
PopupScreen "Tank 1S Status" 480x272
   TextField "Text field_4" at 9,135 size 86x22; Text 'Pressure:'
   IOField "I/O field_1" at 139,130 size 90x25; FormatPattern s999.9; Unit  mBar
      ProcessValue <- "20_TANKS_IP_DATA_RIO_01_THIRD_TANK_TANKS_PRESS"
   TextField "Text field_5" at 9,169 size 113x22; Text 'Water Level:'
   IOField "I/O field_2" at 138,164 size 90x25; FormatPattern 999.9; Unit  %
      ProcessValue <- "20_TANKS_IP_DATA_RIO_01_THIRD_TANK_BWT_LEVEL"
   TextField "Text field_6" at 9,203 size 137x22; Text 'MBG Flow Rate:'
   IOField "I/O field_3" at 139,198 size 90x25; FormatPattern 999.9; Unit  m³/hr
      ProcessValue <- "20_TANKS_IP_DATA_RIO_01_THIRD_TANK_MBG_FLOW"
   TextField "Text field_7" at 9,237 size 135x22; Text 'USD Flow Rate:'
   IOField "I/O field_4" at 139,232 size 90x25; FormatPattern 999.9; Unit  m³/hr
      ProcessValue <- "20_TANKS_IP_DATA_RIO_01_THIRD_TANK_USD_FLOW"
   Button "Button_1" at 50,5 size 191x35; TextOff 'Starboard Tank 1 (1S)'
      on Release: function_efd93a16("Tank 1S Status", 0, 0, -1, 0, 1)
   TextField "Text field_1" at 4,90 size 109x25; Text 'TIME LEFT:'
   GraphicView "Graphic view_1" at 9,46 size 228x32; Picture "Tank Manually Disabled"
   GraphicIOField "Graphic I/O field_1" at 9,46 size 228x32; PictureList "Tank Process Stage_II"
      ProcessValue <- "2100_BTCS_CNTRL_DB_BTCS_STATE"
      Visibility <- "504_Tank Grouping_DB2020_GROUP of TANK 3"
   Button "Button_2" at 4,5 size 45x35; TextOff 'Text'; PictureOff "Graphic_286"
      on Click: function_efd93a16("Tank 1S Status", 0, 0, -1, -1, 1)
   IOField "I/O field_29" at 190,90 size 47x25; FormatPattern 99; Unit m
      ProcessValue <- "504_Tank Grouping_DB2020_Time Left Tank_Time Left m Tank 3"
   IOField "I/O field_8" at 147,90 size 42x25; FormatPattern 99; Unit h
      ProcessValue <- "504_Tank Grouping_DB2020_Time Left Tank_Time Left h Tank 3"
   IOField "I/O field_9" at 104,90 size 42x25; FormatPattern 99; Unit d
      ProcessValue <- "504_Tank Grouping_DB2020_Time Left Tank_Time Left d Tank 3"
   TextField "Text field_8" at 241,134 size 140x22; Text 'Water pH Level:'
   IOField "I/O field_5" at 383,129 size 90x25; FormatPattern 99.9
      ProcessValue <- "20_TANKS_IP_DATA_RIO_01_THIRD_TANK_BWT_PH"
   TextField "Text field_9" at 242,168 size 143x22; Text 'Water DO Level:'
   IOField "I/O field_6" at 383,163 size 90x25; FormatPattern 99.99; Unit  mg/l
      ProcessValue <- "20_TANKS_IP_DATA_RIO_01_THIRD_TANK_BWT_DO"
   TextField "Text field_10" at 241,202 size 174x22; Text 'Water Temperature:'
   IOField "I/O field_7" at 398,197 size 75x25; FormatPattern 999.9; Unit  °C
      ProcessValue <- "20_TANKS_IP_DATA_RIO_01_THIRD_TANK_BWT_TEMP"
   Button "Button_5" at 249,229 size 223x40; TextOff 'Tank Shutdown Alarm'
      Visibility <- "2062_Warning_Data_Alarm Tank S1"
   Button "Button_6" at 248,229 size 224x40; TextOff 'No/Low Water Level'; Authorization "Operate"
      Visibility <- "LT421 1S  TANK LEVEL ALARM_ALARM L"

PopupScreen "Tank 2S Status" 480x272
   TextField "Text field_4" at 4,134 size 86x22; Text 'Pressure:'
   IOField "I/O field_1" at 147,129 size 90x25; FormatPattern s999.9; Unit  mBar
      ProcessValue <- "20_TANKS_IP_DATA_RIO_02_SECOND_TANK_TANKS_PRESS"
   TextField "Text field_5" at 4,168 size 113x22; Text 'Water Level:'
   IOField "I/O field_2" at 147,163 size 90x25; FormatPattern 999.9; Unit  %
      ProcessValue <- "20_TANKS_IP_DATA_RIO_02_SECOND_TANK_BWT_LEVEL"
   TextField "Text field_6" at 4,202 size 137x22; Text 'MBG Flow Rate:'
   IOField "I/O field_3" at 147,197 size 90x25; FormatPattern 999.9; Unit  m³/hr
      ProcessValue <- "20_TANKS_IP_DATA_RIO_02_SECOND_TANK_MBG_FLOW"
   TextField "Text field_7" at 4,236 size 135x22; Text 'USD Flow Rate:'
   IOField "I/O field_4" at 147,231 size 90x25; FormatPattern 999.9; Unit  m³/hr
      ProcessValue <- "20_TANKS_IP_DATA_RIO_02_SECOND_TANK_USD_FLOW"
   Button "Button_1" at 50,5 size 191x35; TextOff 'Starboard Tank 2 (2S)'
      on Release: function_efd93a16("Tank 2S Status", 0, 0, -1, 0, 1)
   TextField "Text field_1" at 5,90 size 109x25; Text 'TIME LEFT:'
   GraphicView "Graphic view_1" at 9,46 size 225x32; Picture "Tank Manually Disabled"
   GraphicIOField "Graphic I/O field_1" at 9,46 size 227x32; PictureList "Tank Process Stage_II"
      ProcessValue <- "2100_BTCS_CNTRL_DB_BTCS_STATE"
      Visibility <- "504_Tank Grouping_DB2020_GROUP of TANK 5"
   Button "Button_2" at 4,5 size 45x35; TextOff 'Text'; PictureOff "Graphic_286"
      on Click: function_efd93a16("Tank 2S Status", 0, 0, -1, -1, 1)
   IOField "I/O field_29" at 189,89 size 47x25; FormatPattern 99; Unit m
      ProcessValue <- "504_Tank Grouping_DB2020_Time Left Tank_Time Left m Tank 5"
   IOField "I/O field_8" at 146,90 size 42x25; FormatPattern 99; Unit h
      ProcessValue <- "504_Tank Grouping_DB2020_Time Left Tank_Time Left h Tank 5"
   IOField "I/O field_9" at 103,90 size 42x25; FormatPattern 99; Unit d
      ProcessValue <- "504_Tank Grouping_DB2020_Time Left Tank_Time Left d Tank 5"
   TextField "Text field_8" at 243,133 size 140x22; Text 'Water pH Level:'
   IOField "I/O field_5" at 382,128 size 90x25; FormatPattern 99.9
      ProcessValue <- "20_TANKS_IP_DATA_RIO_02_SECOND_TANK_BWT_PH"
   TextField "Text field_9" at 243,167 size 143x22; Text 'Water DO Level:'
   IOField "I/O field_6" at 382,162 size 90x25; FormatPattern 99.99; Unit  mg/l
      ProcessValue <- "20_TANKS_IP_DATA_RIO_02_SECOND_TANK_BWT_DO"
   TextField "Text field_10" at 243,201 size 174x22; Text 'Water Temperature:'
   IOField "I/O field_7" at 397,196 size 75x25; FormatPattern 999.9; Unit  °C
      ProcessValue <- "20_TANKS_IP_DATA_RIO_02_SECOND_TANK_BWT_TEMP"
   Group "Group" at 245,228 size 227x40
   Button "Button_5" at 245,228 size 227x40; TextOff 'Tank Shutdown Alarm'
      Visibility <- "2062_Warning_Data_Alarm Tank S2"
   Button "Button_6" at 245,228 size 227x40; TextOff 'No/Low Water Level'; Authorization "Operate"
      Visibility <- "LT421 2S  TANK LEVEL ALARM_ALARM L"

PopupScreen "Tank 2P Status" 480x272
   TextField "Text field_4" at 8,135 size 86x22; Text 'Pressure:'
   IOField "I/O field_1" at 139,130 size 90x25; FormatPattern s999.9; Unit  mBar
      ProcessValue <- "20_TANKS_IP_DATA_RIO_02_FIRST_TANK_TANKS_PRESS"
   TextField "Text field_5" at 8,169 size 113x22; Text 'Water Level:'
   IOField "I/O field_2" at 139,164 size 90x25; FormatPattern 999.9; Unit  %
      ProcessValue <- "20_TANKS_IP_DATA_RIO_02_FIRST_TANK_BWT_LEVEL"
   TextField "Text field_6" at 8,203 size 137x22; Text 'MBG Flow Rate:'
   IOField "I/O field_3" at 139,198 size 90x25; FormatPattern 999.9; Unit  m³/hr
      ProcessValue <- "20_TANKS_IP_DATA_RIO_02_FIRST_TANK_MBG_FLOW"
   TextField "Text field_7" at 8,237 size 135x22; Text 'USD Flow Rate:'
   IOField "I/O field_4" at 139,232 size 90x25; FormatPattern 999.9; Unit  m³/hr
      ProcessValue <- "20_TANKS_IP_DATA_RIO_02_FIRST_TANK_USD_FLOW"
   Button "Button_1" at 51,5 size 188x35; TextOff 'Port Tank 2 (2P)'
      on Release: function_efd93a16("Tank 2P Status", 0, 0, -1, 0, 1)
   TextField "Text field_1" at 4,90 size 109x25; Text 'TIME LEFT:'
   GraphicView "Graphic view_1" at 9,46 size 225x32; Picture "Tank Manually Disabled"
   GraphicIOField "Graphic I/O field_1" at 9,46 size 225x32; PictureList "Tank Process Stage_II"
      ProcessValue <- "2100_BTCS_CNTRL_DB_BTCS_STATE"
      Visibility <- "504_Tank Grouping_DB2020_GROUP of TANK 4"
   Button "Button_2" at 4,5 size 45x35; TextOff 'Text'; PictureOff "Graphic_286"
      on Click: function_efd93a16("Tank 2P Status", 0, 0, -1, -1, 1)
   IOField "I/O field_29" at 187,90 size 47x25; FormatPattern 99; Unit m
      ProcessValue <- "504_Tank Grouping_DB2020_Time Left Tank_Time Left m Tank 4"
   IOField "I/O field_8" at 144,90 size 42x25; FormatPattern 99; Unit h
      ProcessValue <- "504_Tank Grouping_DB2020_Time Left Tank_Time Left h Tank 4"
   IOField "I/O field_9" at 101,90 size 42x25; FormatPattern 99; Unit d
      ProcessValue <- "504_Tank Grouping_DB2020_Time Left Tank_Time Left d Tank 4"
   TextField "Text field_8" at 245,135 size 140x22; Text 'Water pH Level:'
   IOField "I/O field_5" at 385,130 size 90x25; FormatPattern 99.9
      ProcessValue <- "20_TANKS_IP_DATA_RIO_02_FIRST_TANK_BWT_PH"
   TextField "Text field_9" at 245,169 size 143x22; Text 'Water DO Level:'
   IOField "I/O field_6" at 385,164 size 90x25; FormatPattern 99.99; Unit  mg/l
      ProcessValue <- "20_TANKS_IP_DATA_RIO_02_FIRST_TANK_BWT_DO"
   TextField "Text field_10" at 245,203 size 174x22; Text 'Water Temperature:'
   IOField "I/O field_7" at 400,198 size 75x25; FormatPattern 999.9; Unit  °C
      ProcessValue <- "20_TANKS_IP_DATA_RIO_02_FIRST_TANK_BWT_TEMP"
   Group "Group" at 244,226 size 230x40
   Button "Button_5" at 244,226 size 230x40; TextOff 'Tank Shutdown Alarm'
      Visibility <- "2062_Warning_Data_Alarm Tank P2"
   Button "Button_6" at 244,226 size 230x40; TextOff 'No/Low Water Level'; Authorization "Operate"
      Visibility <- "FIT418_2P_ALM_ANALOG_DB_ALARM L"

PopupScreen "Tank 3S Status" 480x272
   TextField "Text field_4" at 9,135 size 86x22; Text 'Pressure:'
   IOField "I/O field_1" at 146,130 size 90x25; FormatPattern s999.9; Unit  mBar
      ProcessValue <- "20_TANKS_IP_DATA_RIO_03_SECOND_TANK_TANKS_PRESS"
   TextField "Text field_5" at 9,169 size 113x22; Text 'Water Level:'
   IOField "I/O field_2" at 146,164 size 90x25; FormatPattern 999.9; Unit  %
      ProcessValue <- "20_TANKS_IP_DATA_RIO_03_SECOND_TANK_BWT_LEVEL"
   TextField "Text field_6" at 9,203 size 137x22; Text 'MBG Flow Rate:'
   IOField "I/O field_3" at 146,198 size 90x25; FormatPattern 999.9; Unit  m³/hr
      ProcessValue <- "20_TANKS_IP_DATA_RIO_03_SECOND_TANK_MBG_FLOW"
   TextField "Text field_7" at 9,237 size 135x22; Text 'USD Flow Rate:'
   IOField "I/O field_4" at 146,232 size 90x25; FormatPattern 999.9; Unit  m³/hr
      ProcessValue <- "20_TANKS_IP_DATA_RIO_03_SECOND_TANK_USD_FLOW"
   Button "Button_1" at 51,5 size 189x35; TextOff 'Starboard Tank 3 (3S)'
      on Release: function_efd93a16("Tank 3S Status", 0, 0, -1, 0, 1)
   TextField "Text field_1" at 5,90 size 109x25; Text 'TIME LEFT:'
   GraphicView "Graphic view_1" at 9,46 size 226x32; Picture "Tank Manually Disabled"
   GraphicIOField "Graphic I/O field_1" at 9,46 size 226x32; PictureList "Tank Process Stage_II"
      ProcessValue <- "2100_BTCS_CNTRL_DB_BTCS_STATE"
      Visibility <- "504_Tank Grouping_DB2020_GROUP of TANK 7"
   Button "Button_2" at 4,5 size 45x35; TextOff 'Text'; PictureOff "Graphic_286"
      on Click: function_efd93a16("Tank 3S Status", 0, 0, -1, -1, 1)
   IOField "I/O field_29" at 189,90 size 47x25; FormatPattern 99; Unit m
      ProcessValue <- "504_Tank Grouping_DB2020_Time Left Tank_Time Left m Tank 7"
   IOField "I/O field_8" at 146,90 size 42x25; FormatPattern 99; Unit h
      ProcessValue <- "504_Tank Grouping_DB2020_Time Left Tank_Time Left h Tank 7"
   IOField "I/O field_9" at 103,90 size 42x25; FormatPattern 99; Unit d
      ProcessValue <- "504_Tank Grouping_DB2020_Time Left Tank_Time Left d Tank 7"
   TextField "Text field_8" at 243,135 size 140x22; Text 'Water pH Level:'
   IOField "I/O field_5" at 383,130 size 90x25; FormatPattern 99.9
      ProcessValue <- "20_TANKS_IP_DATA_RIO_03_SECOND_TANK_BWT_PH"
   TextField "Text field_9" at 243,169 size 143x22; Text 'Water DO Level:'
   IOField "I/O field_6" at 383,164 size 90x25; FormatPattern 99.99; Unit  mg/l
      ProcessValue <- "20_TANKS_IP_DATA_RIO_03_SECOND_TANK_BWT_DO"
   TextField "Text field_10" at 243,203 size 174x22; Text 'Water Temperature:'
   IOField "I/O field_7" at 398,198 size 75x25; FormatPattern 999.9; Unit  °C
      ProcessValue <- "20_TANKS_IP_DATA_RIO_03_SECOND_TANK_BWT_TEMP"
   Group "Group" at 243,228 size 230x40
   Button "Button_5" at 243,228 size 230x40; TextOff 'Tank Shutdown Alarm'
      Visibility <- "2062_Warning_Data_Alarm Tank S3"
   Button "Button_6" at 243,228 size 230x40; TextOff 'No/Low Water Level'; Authorization "Operate"
      Visibility <- "LT421 3S  TANK LEVEL ALARM_ALARM L"

PopupScreen "Tank 3P Status" 480x272
   TextField "Text field_4" at 10,135 size 86x22; Text 'Pressure:'
   IOField "I/O field_1" at 148,130 size 90x25; FormatPattern s999.9; Unit  mBar
      ProcessValue <- "20_TANKS_IP_DATA_RIO_03_FIRST_TANK_TANKS_PRESS"
   TextField "Text field_5" at 10,169 size 113x22; Text 'Water Level:'
   IOField "I/O field_2" at 148,164 size 90x25; FormatPattern 999.9; Unit  %
      ProcessValue <- "20_TANKS_IP_DATA_RIO_03_FIRST_TANK_BWT_LEVEL"
   TextField "Text field_6" at 10,203 size 137x22; Text 'MBG Flow Rate:'
   IOField "I/O field_3" at 148,198 size 90x25; FormatPattern 999.9; Unit  m³/hr
      ProcessValue <- "20_TANKS_IP_DATA_RIO_03_FIRST_TANK_MBG_FLOW"
   TextField "Text field_7" at 10,237 size 135x22; Text 'USD Flow Rate:'
   IOField "I/O field_4" at 148,232 size 90x25; FormatPattern 999.9; Unit  m³/hr
      ProcessValue <- "20_TANKS_IP_DATA_RIO_03_FIRST_TANK_USD_FLOW"
   Button "Button_1" at 51,5 size 191x35; TextOff 'Port Tank 3 (3P)'
      on Release: function_efd93a16("Tank 3P Status", 0, 0, -1, 0, 1)
   TextField "Text field_1" at 6,90 size 109x25; Text 'TIME LEFT:'
   GraphicView "Graphic view_1" at 9,46 size 228x32; Picture "Tank Manually Disabled"
   GraphicIOField "Graphic I/O field_1" at 9,46 size 228x32; PictureList "Tank Process Stage_II"
      ProcessValue <- "2100_BTCS_CNTRL_DB_BTCS_STATE"
      Visibility <- "504_Tank Grouping_DB2020_GROUP of TANK 6"
   Button "Button_2" at 4,5 size 45x35; TextOff 'Text'; PictureOff "Graphic_286"
      on Click: function_efd93a16("Tank 3P Status", 0, 0, -1, -1, 1)
   IOField "I/O field_29" at 190,90 size 47x25; FormatPattern 99; Unit m
      ProcessValue <- "504_Tank Grouping_DB2020_Time Left Tank_Time Left m Tank 6"
   IOField "I/O field_8" at 147,90 size 42x25; FormatPattern 99; Unit h
      ProcessValue <- "504_Tank Grouping_DB2020_Time Left Tank_Time Left h Tank 6"
   IOField "I/O field_9" at 104,90 size 42x25; FormatPattern 99; Unit d
      ProcessValue <- "504_Tank Grouping_DB2020_Time Left Tank_Time Left d Tank 6"
   TextField "Text field_8" at 244,135 size 140x22; Text 'Water pH Level:'
   IOField "I/O field_5" at 383,130 size 90x25; FormatPattern 99.9
      ProcessValue <- "20_TANKS_IP_DATA_RIO_03_FIRST_TANK_BWT_PH"
   TextField "Text field_9" at 244,169 size 143x22; Text 'Water DO Level:'
   IOField "I/O field_6" at 383,164 size 90x25; FormatPattern 99.99; Unit  mg/l
      ProcessValue <- "20_TANKS_IP_DATA_RIO_03_FIRST_TANK_BWT_DO"
   TextField "Text field_10" at 244,203 size 174x22; Text 'Water Temperature:'
   IOField "I/O field_7" at 398,198 size 75x25; FormatPattern 999.9; Unit  °C
      ProcessValue <- "20_TANKS_IP_DATA_RIO_03_FIRST_TANK_BWT_TEMP"
   Group "Group" at 247,227 size 226x40
   Button "Button_5" at 247,227 size 226x40; TextOff 'Tank Shutdown Alarm'
      Visibility <- "2062_Warning_Data_Alarm Tank P3"
   Button "Button_6" at 247,227 size 226x40; TextOff 'No/Low Water Level'; Authorization "Operate"
      Visibility <- "LT422 3P  TANK LEVEL ALARM_ALARM L"

PopupScreen "Tank 4S Status" 480x272
   TextField "Text field_4" at 9,135 size 86x22; Text 'Pressure:'
   IOField "I/O field_1" at 147,130 size 90x25; FormatPattern s999.9; Unit  mBar
      ProcessValue <- "20_TANKS_IP_DATA_RIO_04_SECOND_TANK_TANKS_PRESS"
   TextField "Text field_5" at 9,169 size 113x22; Text 'Water Level:'
   IOField "I/O field_2" at 147,164 size 90x25; FormatPattern 999.9; Unit  %
      ProcessValue <- "20_TANKS_IP_DATA_RIO_04_SECOND_TANK_BWT_LEVEL"
   TextField "Text field_6" at 9,203 size 137x22; Text 'MBG Flow Rate:'
   IOField "I/O field_3" at 147,198 size 90x25; FormatPattern 999.9; Unit  m³/hr
      ProcessValue <- "20_TANKS_IP_DATA_RIO_04_SECOND_TANK_MBG_FLOW"
   TextField "Text field_7" at 9,237 size 135x22; Text 'USD Flow Rate:'
   IOField "I/O field_4" at 147,232 size 90x25; FormatPattern 999.9; Unit  m³/hr
      ProcessValue <- "20_TANKS_IP_DATA_RIO_04_SECOND_TANK_USD_FLOW"
   Button "Button_1" at 50,5 size 191x35; TextOff 'Starboard Tank 4 (4S)'
      on Release: function_efd93a16("Tank 4S Status", 0, 0, -1, 2, 1)
   TextField "Text field_1" at 5,90 size 109x25; Text 'TIME LEFT:'
   GraphicView "Graphic view_1" at 9,46 size 227x32; Picture "Tank Manually Disabled"
   GraphicIOField "Graphic I/O field_1" at 9,46 size 227x32; PictureList "Tank Process Stage_II"
      ProcessValue <- "2100_BTCS_CNTRL_DB_BTCS_STATE"
      Visibility <- "504_Tank Grouping_DB2020_GROUP of TANK 9"
   Button "Button_2" at 4,5 size 45x35; TextOff 'Text'; PictureOff "Graphic_286"
      on Click: function_efd93a16("Tank 4S Status", 0, 0, -1, -1, 1)
   IOField "I/O field_29" at 189,90 size 47x25; FormatPattern 99; Unit m
      ProcessValue <- "504_Tank Grouping_DB2020_Time Left Tank_Time Left m Tank 9"
   IOField "I/O field_8" at 146,90 size 42x25; FormatPattern 99; Unit h
      ProcessValue <- "504_Tank Grouping_DB2020_Time Left Tank_Time Left h Tank 9"
   IOField "I/O field_9" at 103,90 size 42x25; FormatPattern 99; Unit d
      ProcessValue <- "504_Tank Grouping_DB2020_Time Left Tank_Time Left d Tank 9"
   TextField "Text field_8" at 243,135 size 140x22; Text 'Water pH Level:'
   IOField "I/O field_5" at 383,130 size 90x25; FormatPattern 99.9
      ProcessValue <- "20_TANKS_IP_DATA_RIO_04_SECOND_TANK_BWT_PH"
   TextField "Text field_9" at 243,169 size 143x22; Text 'Water DO Level:'
   IOField "I/O field_6" at 383,164 size 90x25; FormatPattern 99.99; Unit  mg/l
      ProcessValue <- "20_TANKS_IP_DATA_RIO_04_SECOND_TANK_BWT_DO"
   TextField "Text field_10" at 243,203 size 174x22; Text 'Water Temperature:'
   IOField "I/O field_7" at 398,198 size 75x25; FormatPattern 999.9; Unit  °C
      ProcessValue <- "20_TANKS_IP_DATA_RIO_04_SECOND_TANK_BWT_TEMP"
   Group "Group" at 243,227 size 230x40
   Button "Button_5" at 243,227 size 230x40; TextOff 'Tank Shutdown Alarm'
      Visibility <- "2062_Warning_Data_Alarm Tank S4"
   Button "Button_6" at 243,227 size 230x40; TextOff 'No/Low Water Level'; Authorization "Operate"
      Visibility <- "LT421 4S  TANK LEVEL ALARM_ALARM L"

PopupScreen "Tank 4P Status" 480x272
   TextField "Text field_4" at 9,135 size 86x22; Text 'Pressure:'
   IOField "I/O field_1" at 148,130 size 90x25; FormatPattern s999.9; Unit  mBar
      ProcessValue <- "20_TANKS_IP_DATA_RIO_04_FIRST_TANK_TANKS_PRESS"
   TextField "Text field_5" at 9,169 size 113x22; Text 'Water Level:'
   IOField "I/O field_2" at 148,164 size 90x25; FormatPattern 999.9; Unit  %
      ProcessValue <- "20_TANKS_IP_DATA_RIO_04_FIRST_TANK_BWT_LEVEL"
   TextField "Text field_6" at 9,203 size 137x22; Text 'MBG Flow Rate:'
   IOField "I/O field_3" at 148,198 size 90x25; FormatPattern 999.9; Unit  m³/hr
      ProcessValue <- "20_TANKS_IP_DATA_RIO_04_FIRST_TANK_MBG_FLOW"
   TextField "Text field_7" at 9,237 size 135x22; Text 'USD Flow Rate:'
   IOField "I/O field_4" at 148,232 size 90x25; FormatPattern 999.9; Unit  m³/hr
      ProcessValue <- "20_TANKS_IP_DATA_RIO_04_FIRST_TANK_USD_FLOW"
   Button "Button_1" at 51,5 size 191x35; TextOff 'Port Tank 4 (4P)'
      on Release: function_efd93a16("Tank 4P Status", 0, 0, -1, 2, 1)
   TextField "Text field_1" at 5,90 size 109x25; Text 'TIME LEFT:'
   GraphicView "Graphic view_1" at 9,46 size 227x32; Picture "Tank Manually Disabled"
   GraphicIOField "Graphic I/O field_1" at 9,46 size 228x32; PictureList "Tank Process Stage_II"
      ProcessValue <- "2100_BTCS_CNTRL_DB_BTCS_STATE"
      Visibility <- "504_Tank Grouping_DB2020_GROUP of TANK 8"
   Button "Button_2" at 4,5 size 45x35; TextOff 'Text'; PictureOff "Graphic_286"
      on Click: function_efd93a16("Tank 4P Status", 0, 0, -1, -1, 1)
   IOField "I/O field_29" at 190,90 size 47x25; FormatPattern 99; Unit m
      ProcessValue <- "504_Tank Grouping_DB2020_Time Left Tank_Time Left m Tank 8"
   IOField "I/O field_8" at 147,90 size 42x25; FormatPattern 99; Unit h
      ProcessValue <- "504_Tank Grouping_DB2020_Time Left Tank_Time Left h Tank 8"
   IOField "I/O field_9" at 104,90 size 42x25; FormatPattern 99; Unit d
      ProcessValue <- "504_Tank Grouping_DB2020_Time Left Tank_Time Left d Tank 8"
   TextField "Text field_8" at 244,135 size 140x22; Text 'Water pH Level:'
   IOField "I/O field_5" at 384,130 size 90x25; FormatPattern 99.9
      ProcessValue <- "20_TANKS_IP_DATA_RIO_04_FIRST_TANK_BWT_PH"
   TextField "Text field_9" at 244,169 size 143x22; Text 'Water DO Level:'
   IOField "I/O field_6" at 384,164 size 90x25; FormatPattern 99.99; Unit  mg/l
      ProcessValue <- "20_TANKS_IP_DATA_RIO_04_FIRST_TANK_BWT_DO"
   TextField "Text field_10" at 244,203 size 174x22; Text 'Water Temperature:'
   IOField "I/O field_7" at 399,198 size 75x25; FormatPattern 999.9; Unit  °C
      ProcessValue <- "20_TANKS_IP_DATA_RIO_04_FIRST_TANK_BWT_TEMP"
   Group "Group" at 244,227 size 230x40
   Button "Button_5" at 244,227 size 230x40; TextOff 'Tank Shutdown Alarm'
      Visibility <- "2062_Warning_Data_Alarm Tank P4"
   Button "Button_6" at 244,227 size 230x40; TextOff 'No/Low Water Level'; Authorization "Operate"
      Visibility <- "LT422 4P  TANK LEVEL ALARM_ALARM L"

PopupScreen "Tank 5S Status" 480x272
   TextField "Text field_4" at 9,135 size 86x22; Text 'Pressure:'
   IOField "I/O field_1" at 147,130 size 90x25; FormatPattern s999.9; Unit  mBar
      ProcessValue <- "20_TANKS_IP_DATA_RIO_05_SECOND_TANK_TANKS_PRESS"
   TextField "Text field_5" at 9,169 size 113x22; Text 'Water Level:'
   IOField "I/O field_2" at 147,164 size 90x25; FormatPattern 999.9; Unit  %
      ProcessValue <- "20_TANKS_IP_DATA_RIO_05_SECOND_TANK_BWT_LEVEL"
   TextField "Text field_6" at 9,203 size 137x22; Text 'MBG Flow Rate:'
   IOField "I/O field_3" at 147,198 size 90x25; FormatPattern 999.9; Unit  m³/hr
      ProcessValue <- "20_TANKS_IP_DATA_RIO_05_SECOND_TANK_MBG_FLOW"
   TextField "Text field_7" at 9,237 size 135x22; Text 'USD Flow Rate:'
   IOField "I/O field_4" at 147,232 size 90x25; FormatPattern 999.9; Unit  m³/hr
      ProcessValue <- "20_TANKS_IP_DATA_RIO_05_SECOND_TANK_USD_FLOW"
   Button "Button_1" at 50,5 size 192x35; TextOff 'Starboard Tank 5 (5S)'
      on Release: function_efd93a16("Tank 5S Status", 0, 0, -1, 2, 1)
   TextField "Text field_1" at 6,90 size 109x25; Text 'TIME LEFT:'
   GraphicView "Graphic view_1" at 9,46 size 228x32; Picture "Tank Manually Disabled"
   GraphicIOField "Graphic I/O field_1" at 9,46 size 228x32; PictureList "Tank Process Stage_II"
      ProcessValue <- "2100_BTCS_CNTRL_DB_BTCS_STATE"
      Visibility <- "504_Tank Grouping_DB2020_GROUP of TANK 11"
   Button "Button_2" at 4,5 size 45x35; TextOff 'Text'; PictureOff "Graphic_286"
      on Click: function_efd93a16("Tank 5S Status", 0, 0, -1, -1, 1)
   IOField "I/O field_29" at 190,90 size 47x25; FormatPattern 99; Unit m
      ProcessValue <- "504_Tank Grouping_DB2020_Time Left Tank_Time Left m Tank 11"
   IOField "I/O field_8" at 147,90 size 42x25; FormatPattern 99; Unit h
      ProcessValue <- "504_Tank Grouping_DB2020_Time Left Tank_Time Left h Tank 11"
   IOField "I/O field_9" at 104,90 size 42x25; FormatPattern 99; Unit d
      ProcessValue <- "504_Tank Grouping_DB2020_Time Left Tank_Time Left d Tank 11"
   TextField "Text field_8" at 243,135 size 140x22; Text 'Water pH Level:'
   IOField "I/O field_5" at 383,130 size 90x25; FormatPattern 99.9
      ProcessValue <- "20_TANKS_IP_DATA_RIO_05_SECOND_TANK_BWT_PH"
   TextField "Text field_9" at 243,169 size 143x22; Text 'Water DO Level:'
   IOField "I/O field_6" at 383,164 size 90x25; FormatPattern 99.99; Unit  mg/l
      ProcessValue <- "20_TANKS_IP_DATA_RIO_05_SECOND_TANK_BWT_DO"
   TextField "Text field_10" at 243,203 size 174x22; Text 'Water Temperature:'
   IOField "I/O field_7" at 398,198 size 75x25; FormatPattern 999.9; Unit  °C
      ProcessValue <- "20_TANKS_IP_DATA_RIO_05_SECOND_TANK_BWT_TEMP"
   Group "Group" at 245,227 size 228x40
   Button "Button_5" at 245,227 size 228x40; TextOff 'Tank Shutdown Alarm'
      Visibility <- "2062_Warning_Data_Alarm Tank S5"
   Button "Button_6" at 245,227 size 228x40; TextOff 'No/Low Water Level'; Authorization "Operate"
      Visibility <- "LT421 5S  TANK LEVEL ALARM_ALARM L"

PopupScreen "Tank 5P Status" 480x272
   TextField "Text field_4" at 9,135 size 86x22; Text 'Pressure:'
   IOField "I/O field_1" at 150,130 size 90x25; FormatPattern s999.9; Unit  mBar
      ProcessValue <- "20_TANKS_IP_DATA_RIO_05_FIRST_TANK_TANKS_PRESS"
   TextField "Text field_5" at 9,169 size 113x22; Text 'Water Level:'
   IOField "I/O field_2" at 150,164 size 90x25; FormatPattern 999.9; Unit  %
      ProcessValue <- "20_TANKS_IP_DATA_RIO_05_FIRST_TANK_BWT_LEVEL"
   TextField "Text field_6" at 9,203 size 137x22; Text 'MBG Flow Rate:'
   IOField "I/O field_3" at 150,198 size 90x25; FormatPattern 999.9; Unit  m³/hr
      ProcessValue <- "20_TANKS_IP_DATA_RIO_05_FIRST_TANK_MBG_FLOW"
   TextField "Text field_7" at 9,237 size 135x22; Text 'USD Flow Rate:'
   IOField "I/O field_4" at 150,232 size 90x25; FormatPattern 999.9; Unit  m³/hr
      ProcessValue <- "20_TANKS_IP_DATA_RIO_05_FIRST_TANK_USD_FLOW"
   Button "Button_1" at 51,5 size 194x35; TextOff 'Port Tank 5 (5P)'
      on Release: function_efd93a16("Tank 5P Status", 0, 0, -1, 2, 1)
   TextField "Text field_1" at 5,90 size 109x25; Text 'TIME LEFT:'
   GraphicView "Graphic view_1" at 9,46 size 231x32; Picture "Tank Manually Disabled"
   GraphicIOField "Graphic I/O field_1" at 9,46 size 231x32; PictureList "Tank Process Stage_II"
      ProcessValue <- "2100_BTCS_CNTRL_DB_BTCS_STATE"
      Visibility <- "504_Tank Grouping_DB2020_GROUP of TANK 10"
   Button "Button_2" at 4,5 size 45x35; TextOff 'Text'; PictureOff "Graphic_286"
      on Click: function_efd93a16("Tank 5P Status", 0, 0, -1, -1, 1)
   IOField "I/O field_29" at 193,90 size 47x25; FormatPattern 99; Unit m
      ProcessValue <- "504_Tank Grouping_DB2020_Time Left Tank_Time Left m Tank 10"
   IOField "I/O field_8" at 148,90 size 42x25; FormatPattern 99; Unit h
      ProcessValue <- "504_Tank Grouping_DB2020_Time Left Tank_Time Left h Tank 10"
   IOField "I/O field_9" at 103,90 size 42x25; FormatPattern 99; Unit d
      ProcessValue <- "504_Tank Grouping_DB2020_Time Left Tank_Time Left d Tank 10"
   TextField "Text field_8" at 244,135 size 140x22; Text 'Water pH Level:'
   IOField "I/O field_5" at 384,130 size 90x25; FormatPattern 99.9
      ProcessValue <- "20_TANKS_IP_DATA_RIO_05_FIRST_TANK_BWT_PH"
   TextField "Text field_9" at 244,169 size 143x22; Text 'Water DO Level:'
   IOField "I/O field_6" at 384,164 size 90x25; FormatPattern 99.99; Unit  mg/l
      ProcessValue <- "20_TANKS_IP_DATA_RIO_05_FIRST_TANK_BWT_DO"
   TextField "Text field_10" at 244,203 size 174x22; Text 'Water Temperature:'
   IOField "I/O field_7" at 399,198 size 75x25; FormatPattern 999.9; Unit  °C
      ProcessValue <- "20_TANKS_IP_DATA_RIO_05_FIRST_TANK_BWT_TEMP"
   Group "Group" at 247,228 size 227x40
   Button "Button_5" at 247,228 size 227x40; TextOff 'Tank Shutdown Alarm'
      Visibility <- "2062_Warning_Data_Alarm Tank P5"
   Button "Button_6" at 247,228 size 227x40; TextOff 'No/Low Water Level'; Authorization "Operate"
      Visibility <- "LT422 5P  TANK LEVEL ALARM_ALARM L"

